screen "Parametry proc. i awarie" 800x434
   TextField "Text field_1" at 141,0 size 176x23; Text 'Parametry procesu'
   IOField "I/O field_1" at 19,64 size 85x25; FormatPattern 999.9
      ProcessValue <- "HMI komunikacja_HMI poziom cieczy Z1"
   TextField "Text field_2" at 560,0 size 142x23; Text 'Zasilanie pomp'
   TextField "Text field_3" at 36,23 size 89x21; Text 'Zbiornik 1'
   TextField "Text field_4" at 183,23 size 84x21; Text 'Zbiornik 2'
   TextField "Text field_5" at 330,23 size 84x21; Text 'Zbiornik 3'
   TextField "Text field_6" at 183,228 size 84x21; Text 'Zbiornik 4'
   TextField "Text field_7" at 0,103 size 154x18; Text 'Temperatura procesu'
   TextField "Text field_8" at 0,42 size 101x18; Text 'Poziom cieczy'
   TextField "Text field_9" at 148,42 size 101x18; Text 'Poziom cieczy'
   TextField "Text field_10" at 0,163 size 165x18; Text 'Czas utrzymania temp.'
   TextField "Text field_11" at 148,163 size 165x18; Text 'Czas utrzymania temp.'
   TextField "Text field_12" at 148,103 size 154x18; Text 'Temperatura procesu'
   TextField "Text field_13" at 296,42 size 101x18; Text 'Poziom cieczy'
   TextField "Text field_14" at 296,103 size 154x18; Text 'Temperatura procesu'
   TextField "Text field_15" at 296,163 size 165x18; Text 'Czas utrzymania temp.'
   TextField "Text field_16" at 148,248 size 167x18; Text 'Poziom cieczy (1+2+3)'
   TextField "Text field_17" at 148,307 size 154x18; Text 'Temperatura procesu'
   TextField "Text field_18" at 148,367 size 165x18; Text 'Czas utrzymania temp.'
   TextField "Text field_19" at 510,90 size 16x23; Text 'Text'
   TextField "Text field_20" at 681,25 size 67x20; Text 'Pompa 2'
   TextField "Text field_21" at 507,25 size 67x20; Text 'Pompa 1'
   TextField "Text field_22" at 507,125 size 67x20; Text 'Pompa 3'
   TextField "Text field_23" at 681,125 size 67x20; Text 'Pompa 4'
   TextField "Text field_24" at 681,330 size 67x20; Text 'Pompa 8'
   TextField "Text field_25" at 507,228 size 67x20; Text 'Pompa 5'
   TextField "Text field_26" at 507,330 size 67x20; Text 'Pompa 7'
   TextField "Text field_27" at 681,228 size 67x20; Text 'Pompa 6'
   IOField "I/O field_2" at 166,64 size 85x25; FormatPattern 999.9
      ProcessValue <- "HMI komunikacja_HMI poziom cieczy Z2"
   IOField "I/O field_3" at 314,64 size 85x25; FormatPattern 999.9
      ProcessValue <- "HMI komunikacja_HMI poziom cieczy Z3"
   IOField "I/O field_4" at 19,129 size 85x25; FormatPattern 999
      ProcessValue <- "HMI komunikacja_HMI Temp max Z1"
   IOField "I/O field_5" at 19,188 size 85x25; FormatPattern 999
      ProcessValue <- "HMI komunikacja_HMI czas utrz T  Z1"
   IOField "I/O field_6" at 166,128 size 85x25; FormatPattern 999
      ProcessValue <- "HMI komunikacja_HMI Temp max Z2"
   IOField "I/O field_7" at 167,188 size 85x25; FormatPattern 999
      ProcessValue <- "HMI komunikacja_HMI czas utrz T  Z2"
   IOField "I/O field_8" at 314,129 size 85x25; FormatPattern 999
      ProcessValue <- "HMI komunikacja_HMI Temp max Z3"
   IOField "I/O field_9" at 314,187 size 85x25; FormatPattern 999
      ProcessValue <- "HMI komunikacja_HMI czas utrz T  Z3"
   IOField "I/O field_10" at 167,271 size 85x25; FormatPattern 999.9
      ProcessValue <- "HMI komunikacja_HMI poziom cieczy Z4"
   IOField "I/O field_11" at 167,332 size 85x25; FormatPattern 999
      ProcessValue <- "HMI komunikacja_HMI Temp max Z4"
   IOField "I/O field_12" at 167,393 size 85x25; FormatPattern 999
      ProcessValue <- "HMI komunikacja_HMI czas utrz T  Z4"
   Switch "Switch_1" at 485,49 size 103x48; TextOn 'OFF'; CaptionText 'Switch'; TextOff 'ON'
      ProcessValue <- "OPC - do LabVIEW_HMI konserwacja P1"
      Appearance <- "OPC - do LabVIEW_HMI konserwacja P1"
   Switch "Switch_2" at 659,49 size 103x48; TextOn 'OFF'; CaptionText 'Switch'; TextOff 'ON'
      ProcessValue <- "OPC - do LabVIEW_HMI konserwacja P2"
      Appearance <- "OPC - do LabVIEW_HMI konserwacja P2"
   Switch "Switch_3" at 485,152 size 103x48; TextOn 'OFF'; CaptionText 'Switch'; TextOff 'ON'
      ProcessValue <- "OPC - do LabVIEW_HMI konserwacja P3"
      Appearance <- "OPC - do LabVIEW_HMI konserwacja P3"
   Switch "Switch_4" at 485,255 size 103x48; TextOn 'OFF'; CaptionText 'Switch'; TextOff 'ON'
      Appearance <- "OPC - do LabVIEW_HMI konserwacja P5"
      ProcessValue <- "OPC - do LabVIEW_HMI konserwacja P5"
   Switch "Switch_5" at 485,358 size 103x48; TextOn 'OFF'; CaptionText 'Switch'; TextOff 'ON'
      ProcessValue <- "OPC - do LabVIEW_HMI konserwacja P7"
      Appearance <- "OPC - do LabVIEW_HMI konserwacja P7"
   Switch "Switch_6" at 658,156 size 103x48; TextOn 'OFF'; CaptionText 'Switch'; TextOff 'ON'
      ProcessValue <- "OPC - do LabVIEW_HMI konserwacja P4"
      Appearance <- "OPC - do LabVIEW_HMI konserwacja P4"
   Switch "Switch_7" at 659,255 size 103x48; TextOn 'OFF'; CaptionText 'Switch'; TextOff 'ON'
      Appearance <- "OPC - do LabVIEW_HMI konserwacja P6"
      ProcessValue <- "OPC - do LabVIEW_HMI konserwacja P6"
   Switch "Switch_8" at 659,358 size 103x48; TextOn 'OFF'; CaptionText 'Switch'; TextOff 'ON'
      ProcessValue <- "OPC - do LabVIEW_HMI konserwacja P8"
      Appearance <- "OPC - do LabVIEW_HMI konserwacja P8"
   Circle "Circle_1" at 46,297 size 48x48
      Appearance <- "HMI komunikacja_Blokada zmiany par. PRO"
   TextField "Text field_30" at 0,259 size 167x38; Text 'Możliwa zmiana parametrów procesu'

screen "Wykresy" 800x434
   TextField "Text field_1" at 0,0 size 376x22; Text 'Objętość i temperatura cieczy w zbiorniku 1'
   TextField "Text field_2" at 400,0 size 376x22; Text 'Objętość i temperatura cieczy w zbiorniku 2'
   TextField "Text field_3" at 0,215 size 376x22; Text 'Objętość i temperatura cieczy w zbiorniku 3'
   TextField "Text field_5" at 400,215 size 376x22; Text 'Objętość i temperatura cieczy w zbiorniku 4'
   Button "Button_1" at 104,31 size 192x32; TextOff 'Wykres Zbiornik 1'
      on Click: ActivateScreen("Wykres Zbiornik 1", 0)
   Button "Button_2" at 504,31 size 192x32; TextOff 'Wykres Zbiornik 2'
      on Click: ActivateScreen("Wykres Zbiornik 2", 0)
   Button "Button_3" at 104,247 size 192x32; TextOff 'Wykres Zbiornik 3'
      on Click: ActivateScreen("Wykres Zbiornik 3", 0)
   Button "Button_4" at 504,247 size 192x32; TextOff 'Wykres Zbiornik 4'
      on Click: ActivateScreen("Wykres Zbiornik 4", 0)
   TextField "Text field_4" at 1,71 size 168x22; Text 'Temperatura P1-P2'
   TextField "Text field_6" at 1,287 size 168x22; Text 'Temperatura P5-P6'
   TextField "Text field_7" at 400,71 size 168x22; Text 'Temperatura P3-P4'
   TextField "Text field_8" at 400,287 size 168x22; Text 'Temperatura P7-P8'
   Button "Button_5" at 104,101 size 192x32; TextOff 'Temperatura P1-P2'
      on Click: ActivateScreen("Temperatura P1-P2", 0)
   Button "Button_6" at 504,101 size 192x32; TextOff 'Temperatura P3-P4'
      on Click: ActivateScreen("Temperatura P3-P4", 0)
   Button "Button_7" at 104,317 size 192x32; TextOff 'Temperatura P5-P6'
      on Click: ActivateScreen("Temperatura P5-P6", 0)
   Button "Button_8" at 504,317 size 192x32; TextOff 'Temperatura P7-P8'
      on Click: ActivateScreen("Temperatura P7-P8", 0)

screen "Wykres Zbiornik 1" 800x434
   TextField "Text field_1" at 0,0 size 295x17; Text 'Objętość i temperatura cieczy w zbiorniku 1'
   TrendView "Trend view_1" at 3,19 size 792x411

screen "Wykres Zbiornik 2" 800x434
   TextField "Text field_2" at 0,0 size 295x17; Text 'Objętość i temperatura cieczy w zbiorniku 2'
   TrendView "Trend view_2" at 3,19 size 792x411

screen "Wykres Zbiornik 3" 800x434
   TextField "Text field_2" at 0,0 size 295x17; Text 'Objętość i temperatura cieczy w zbiorniku 3'
   TrendView "Trend view_3" at 3,19 size 792x411

screen "Wykres Zbiornik 4" 800x434
   TextField "Text field_2" at 3,2 size 199x17; Text 'Objętość cieczy w zbiorniku 4'
   TrendView "Trend view_4" at 3,19 size 792x411
   TextField "Text field_1" at 597,2 size 199x17; Text 'Temperatura cieczy w zbiorniku 4'

screen "Temperatura P1-P2" 800x434
   TextField "Text field_1" at 0,0 size 133x17; Text 'Temperatura P1-P2'
   TrendView "Trend view_1" at 3,19 size 792x411

screen "Temperatura P3-P4" 800x434
   TextField "Text field_1" at 0,0 size 133x17; Text 'Temperatura P3-P4'
   TrendView "Trend view_1" at 3,19 size 792x411

screen "Temperatura P5-P6" 800x434
   TextField "Text field_1" at 0,0 size 133x17; Text 'Temperatura P5-P6'
   TrendView "Trend view_1" at 3,19 size 792x411

screen "Temperatura P7-P8" 800x434
   TextField "Text field_1" at 0,0 size 133x17; Text 'Temperatura P7-P8'
   TrendView "Trend view_1" at 3,19 size 792x411
*)